REGION Network 15
   // ***************************************************************************************************************************************************
   // 
   // TC MAP SDC OUT Function Block FB118 - Maps Traffic Cop Zone motion Function blocks. Motion commands are determined at the zone position level and indexed by Zone number and stored in 
   //  "DB116_TC_ZoneMotionControl" DB. Block copies Traffic cop motion commands to the respective Carrier trafic cop and stores in TC_SDC_OUT Tag which is indexed by carrier number. 
   // 
   // ***************************************************************************************************************************************************
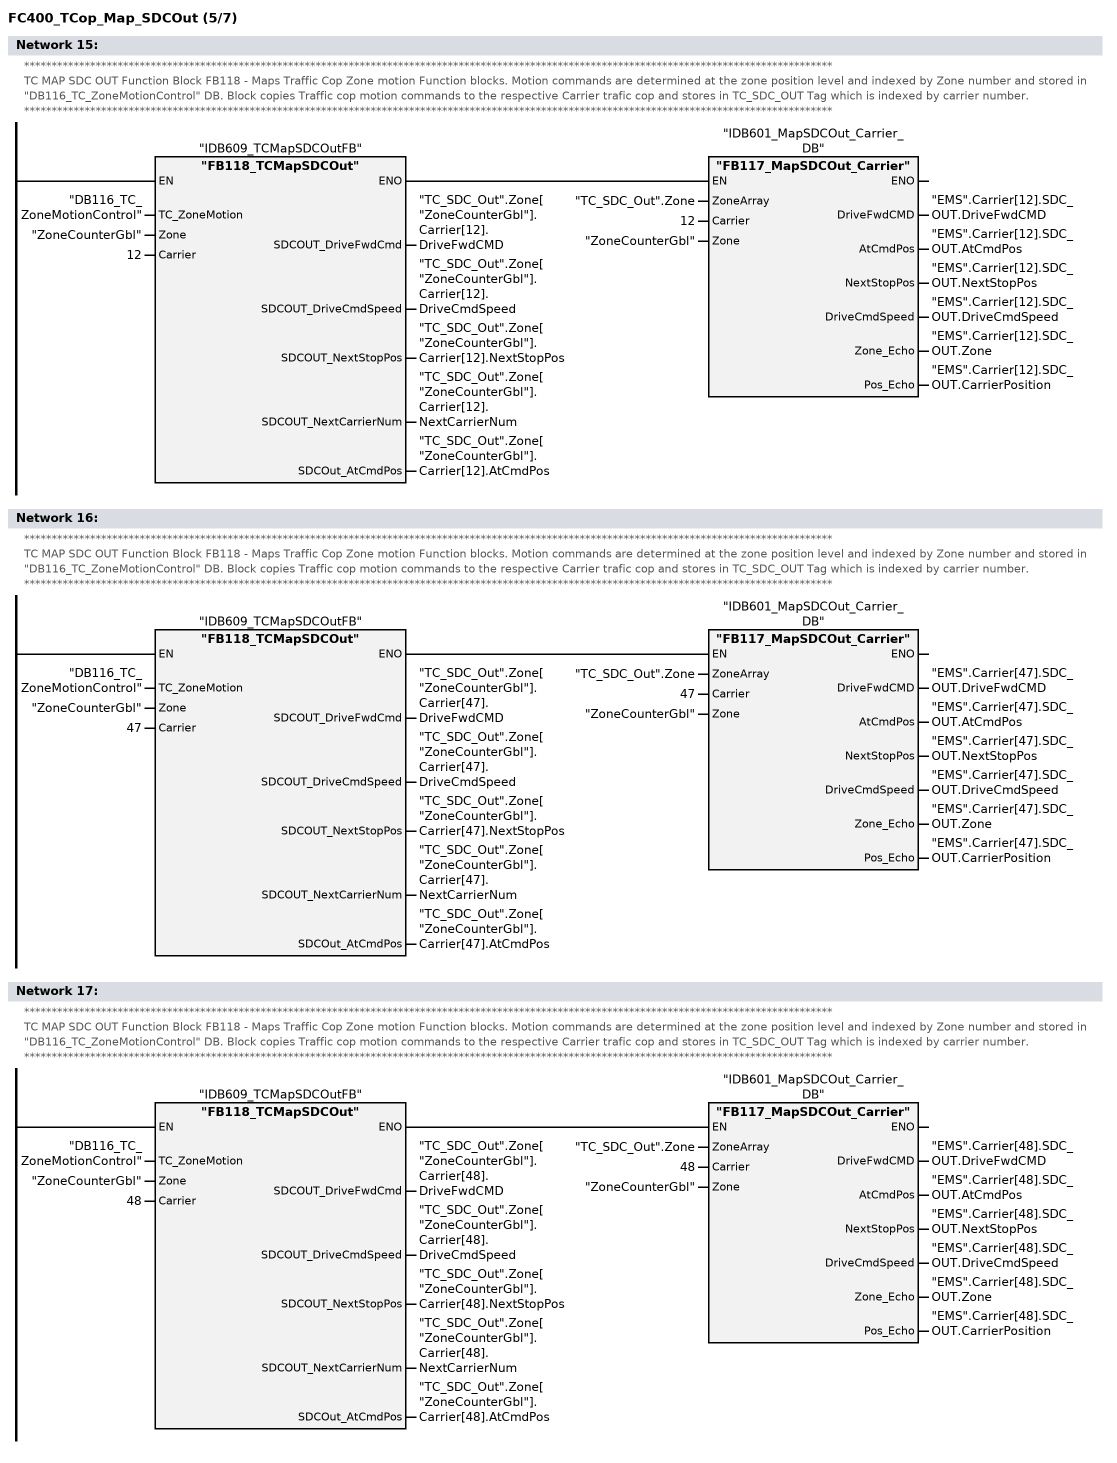
   RUNG wire#powerrail
      "IDB609_TCMapSDCOutFB"(TC_ZoneMotion := "DB116_TC_ZoneMotionControl", Zone := "ZoneCounterGbl", Carrier := 12, SDCOUT_DriveFwdCmd => "TC_SDC_Out".Zone["ZoneCounterGbl"].Carrier[12].DriveFwdCMD, SDCOUT_DriveCmdSpeed => "TC_SDC_Out".Zone["ZoneCounterGbl"].Carrier[12].DriveCmdSpeed, SDCOUT_NextStopPos => "TC_SDC_Out".Zone["ZoneCounterGbl"].Carrier[12].NextStopPos, SDCOUT_NextCarrierNum => "TC_SDC_Out".Zone["ZoneCounterGbl"].Carrier[12].NextCarrierNum, SDCOut_AtCmdPos => "TC_SDC_Out".Zone["ZoneCounterGbl"].Carrier[12].AtCmdPos)
      "IDB601_MapSDCOut_Carrier_DB"(ZoneArray := "TC_SDC_Out".Zone, Carrier := 12, Zone := "ZoneCounterGbl", DriveFwdCMD => "EMS".Carrier[12].SDC_OUT.DriveFwdCMD, AtCmdPos => "EMS".Carrier[12].SDC_OUT.AtCmdPos, NextStopPos => "EMS".Carrier[12].SDC_OUT.NextStopPos, DriveCmdSpeed => "EMS".Carrier[12].SDC_OUT.DriveCmdSpeed, Zone_Echo => "EMS".Carrier[12].SDC_OUT.Zone, Pos_Echo => "EMS".Carrier[12].SDC_OUT.CarrierPosition)
   END_RUNG
   // the same network as SCL:
   "IDB609_TCMapSDCOutFB"(TC_ZoneMotion := "DB116_TC_ZoneMotionControl",   // "FB118_TCMapSDCOut"
                          Zone := "ZoneCounterGbl",
                          Carrier := 12,
                          SDCOUT_DriveFwdCmd => "TC_SDC_Out".Zone["ZoneCounterGbl"].Carrier[12].DriveFwdCMD,
                          SDCOUT_DriveCmdSpeed => "TC_SDC_Out".Zone["ZoneCounterGbl"].Carrier[12].DriveCmdSpeed,
                          SDCOUT_NextStopPos => "TC_SDC_Out".Zone["ZoneCounterGbl"].Carrier[12].NextStopPos,
                          SDCOUT_NextCarrierNum => "TC_SDC_Out".Zone["ZoneCounterGbl"].Carrier[12].NextCarrierNum,
                          SDCOut_AtCmdPos => "TC_SDC_Out".Zone["ZoneCounterGbl"].Carrier[12].AtCmdPos,
                          ENO => #_w1);
   IF #_w1 THEN
       "IDB601_MapSDCOut_Carrier_DB"(ZoneArray := "TC_SDC_Out".Zone,   // "FB117_MapSDCOut_Carrier"
                               Carrier := 12,
                               Zone := "ZoneCounterGbl",
                               DriveFwdCMD => "EMS".Carrier[12].SDC_OUT.DriveFwdCMD,
                               AtCmdPos => "EMS".Carrier[12].SDC_OUT.AtCmdPos,
                               NextStopPos => "EMS".Carrier[12].SDC_OUT.NextStopPos,
                               DriveCmdSpeed => "EMS".Carrier[12].SDC_OUT.DriveCmdSpeed,
                               Zone_Echo => "EMS".Carrier[12].SDC_OUT.Zone,
                               Pos_Echo => "EMS".Carrier[12].SDC_OUT.CarrierPosition);
   END_IF;
END_REGION

REGION Network 16
   // ***************************************************************************************************************************************************
   // 
   // TC MAP SDC OUT Function Block FB118 - Maps Traffic Cop Zone motion Function blocks. Motion commands are determined at the zone position level and indexed by Zone number and stored in 
   //  "DB116_TC_ZoneMotionControl" DB. Block copies Traffic cop motion commands to the respective Carrier trafic cop and stores in TC_SDC_OUT Tag which is indexed by carrier number. 
   // 
   // ***************************************************************************************************************************************************
   RUNG wire#powerrail
      "IDB609_TCMapSDCOutFB"(TC_ZoneMotion := "DB116_TC_ZoneMotionControl", Zone := "ZoneCounterGbl", Carrier := 47, SDCOUT_DriveFwdCmd => "TC_SDC_Out".Zone["ZoneCounterGbl"].Carrier[47].DriveFwdCMD, SDCOUT_DriveCmdSpeed => "TC_SDC_Out".Zone["ZoneCounterGbl"].Carrier[47].DriveCmdSpeed, SDCOUT_NextStopPos => "TC_SDC_Out".Zone["ZoneCounterGbl"].Carrier[47].NextStopPos, SDCOUT_NextCarrierNum => "TC_SDC_Out".Zone["ZoneCounterGbl"].Carrier[47].NextCarrierNum, SDCOut_AtCmdPos => "TC_SDC_Out".Zone["ZoneCounterGbl"].Carrier[47].AtCmdPos)
      "IDB601_MapSDCOut_Carrier_DB"(ZoneArray := "TC_SDC_Out".Zone, Carrier := 47, Zone := "ZoneCounterGbl", DriveFwdCMD => "EMS".Carrier[47].SDC_OUT.DriveFwdCMD, AtCmdPos => "EMS".Carrier[47].SDC_OUT.AtCmdPos, NextStopPos => "EMS".Carrier[47].SDC_OUT.NextStopPos, DriveCmdSpeed => "EMS".Carrier[47].SDC_OUT.DriveCmdSpeed, Zone_Echo => "EMS".Carrier[47].SDC_OUT.Zone, Pos_Echo => "EMS".Carrier[47].SDC_OUT.CarrierPosition)
   END_RUNG
   // the same network as SCL:
   "IDB609_TCMapSDCOutFB"(TC_ZoneMotion := "DB116_TC_ZoneMotionControl",   // "FB118_TCMapSDCOut"
                          Zone := "ZoneCounterGbl",
                          Carrier := 47,
                          SDCOUT_DriveFwdCmd => "TC_SDC_Out".Zone["ZoneCounterGbl"].Carrier[47].DriveFwdCMD,
                          SDCOUT_DriveCmdSpeed => "TC_SDC_Out".Zone["ZoneCounterGbl"].Carrier[47].DriveCmdSpeed,
                          SDCOUT_NextStopPos => "TC_SDC_Out".Zone["ZoneCounterGbl"].Carrier[47].NextStopPos,
                          SDCOUT_NextCarrierNum => "TC_SDC_Out".Zone["ZoneCounterGbl"].Carrier[47].NextCarrierNum,
                          SDCOut_AtCmdPos => "TC_SDC_Out".Zone["ZoneCounterGbl"].Carrier[47].AtCmdPos,
                          ENO => #_w1);
   IF #_w1 THEN
       "IDB601_MapSDCOut_Carrier_DB"(ZoneArray := "TC_SDC_Out".Zone,   // "FB117_MapSDCOut_Carrier"
                               Carrier := 47,
                               Zone := "ZoneCounterGbl",
                               DriveFwdCMD => "EMS".Carrier[47].SDC_OUT.DriveFwdCMD,
                               AtCmdPos => "EMS".Carrier[47].SDC_OUT.AtCmdPos,
                               NextStopPos => "EMS".Carrier[47].SDC_OUT.NextStopPos,
                               DriveCmdSpeed => "EMS".Carrier[47].SDC_OUT.DriveCmdSpeed,
                               Zone_Echo => "EMS".Carrier[47].SDC_OUT.Zone,
                               Pos_Echo => "EMS".Carrier[47].SDC_OUT.CarrierPosition);
   END_IF;
END_REGION

REGION Network 17
   // ***************************************************************************************************************************************************
   // 
   // TC MAP SDC OUT Function Block FB118 - Maps Traffic Cop Zone motion Function blocks. Motion commands are determined at the zone position level and indexed by Zone number and stored in 
   //  "DB116_TC_ZoneMotionControl" DB. Block copies Traffic cop motion commands to the respective Carrier trafic cop and stores in TC_SDC_OUT Tag which is indexed by carrier number. 
   // 
   // ***************************************************************************************************************************************************
   RUNG wire#powerrail
      "IDB609_TCMapSDCOutFB"(TC_ZoneMotion := "DB116_TC_ZoneMotionControl", Zone := "ZoneCounterGbl", Carrier := 48, SDCOUT_DriveFwdCmd => "TC_SDC_Out".Zone["ZoneCounterGbl"].Carrier[48].DriveFwdCMD, SDCOUT_DriveCmdSpeed => "TC_SDC_Out".Zone["ZoneCounterGbl"].Carrier[48].DriveCmdSpeed, SDCOUT_NextStopPos => "TC_SDC_Out".Zone["ZoneCounterGbl"].Carrier[48].NextStopPos, SDCOUT_NextCarrierNum => "TC_SDC_Out".Zone["ZoneCounterGbl"].Carrier[48].NextCarrierNum, SDCOut_AtCmdPos => "TC_SDC_Out".Zone["ZoneCounterGbl"].Carrier[48].AtCmdPos)
      "IDB601_MapSDCOut_Carrier_DB"(ZoneArray := "TC_SDC_Out".Zone, Carrier := 48, Zone := "ZoneCounterGbl", DriveFwdCMD => "EMS".Carrier[48].SDC_OUT.DriveFwdCMD, AtCmdPos => "EMS".Carrier[48].SDC_OUT.AtCmdPos, NextStopPos => "EMS".Carrier[48].SDC_OUT.NextStopPos, DriveCmdSpeed => "EMS".Carrier[48].SDC_OUT.DriveCmdSpeed, Zone_Echo => "EMS".Carrier[48].SDC_OUT.Zone, Pos_Echo => "EMS".Carrier[48].SDC_OUT.CarrierPosition)
   END_RUNG
   // the same network as SCL:
   "IDB609_TCMapSDCOutFB"(TC_ZoneMotion := "DB116_TC_ZoneMotionControl",   // "FB118_TCMapSDCOut"
                          Zone := "ZoneCounterGbl",
                          Carrier := 48,
                          SDCOUT_DriveFwdCmd => "TC_SDC_Out".Zone["ZoneCounterGbl"].Carrier[48].DriveFwdCMD,
                          SDCOUT_DriveCmdSpeed => "TC_SDC_Out".Zone["ZoneCounterGbl"].Carrier[48].DriveCmdSpeed,
                          SDCOUT_NextStopPos => "TC_SDC_Out".Zone["ZoneCounterGbl"].Carrier[48].NextStopPos,
                          SDCOUT_NextCarrierNum => "TC_SDC_Out".Zone["ZoneCounterGbl"].Carrier[48].NextCarrierNum,
                          SDCOut_AtCmdPos => "TC_SDC_Out".Zone["ZoneCounterGbl"].Carrier[48].AtCmdPos,
                          ENO => #_w1);
   IF #_w1 THEN
       "IDB601_MapSDCOut_Carrier_DB"(ZoneArray := "TC_SDC_Out".Zone,   // "FB117_MapSDCOut_Carrier"
                               Carrier := 48,
                               Zone := "ZoneCounterGbl",
                               DriveFwdCMD => "EMS".Carrier[48].SDC_OUT.DriveFwdCMD,
                               AtCmdPos => "EMS".Carrier[48].SDC_OUT.AtCmdPos,
                               NextStopPos => "EMS".Carrier[48].SDC_OUT.NextStopPos,
                               DriveCmdSpeed => "EMS".Carrier[48].SDC_OUT.DriveCmdSpeed,
                               Zone_Echo => "EMS".Carrier[48].SDC_OUT.Zone,
                               Pos_Echo => "EMS".Carrier[48].SDC_OUT.CarrierPosition);
   END_IF;
END_REGION

REGION Network 18
   // ***************************************************************************************************************************************************
   // 
   // TC MAP SDC OUT Function Block FB118 - Maps Traffic Cop Zone motion Function blocks. Motion commands are determined at the zone position level and indexed by Zone number and stored in 
   //  "DB116_TC_ZoneMotionControl" DB. Block copies Traffic cop motion commands to the respective Carrier trafic cop and stores in TC_SDC_OUT Tag which is indexed by carrier number. 
   // 
   // ***************************************************************************************************************************************************
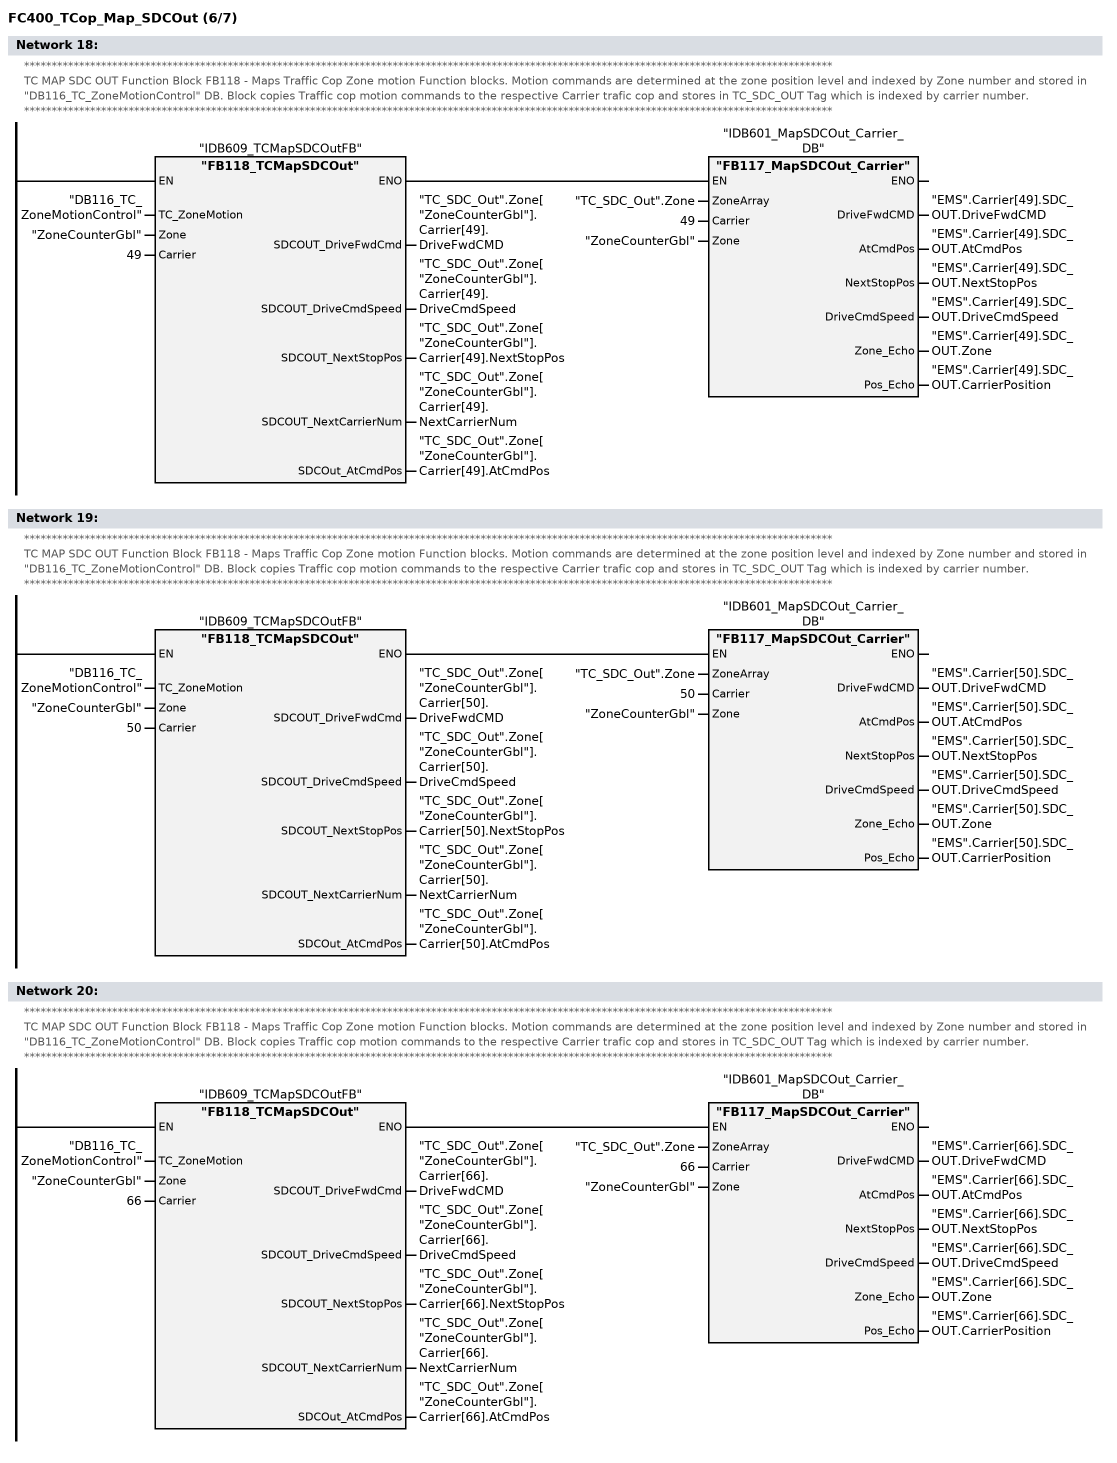
   RUNG wire#powerrail
      "IDB609_TCMapSDCOutFB"(TC_ZoneMotion := "DB116_TC_ZoneMotionControl", Zone := "ZoneCounterGbl", Carrier := 49, SDCOUT_DriveFwdCmd => "TC_SDC_Out".Zone["ZoneCounterGbl"].Carrier[49].DriveFwdCMD, SDCOUT_DriveCmdSpeed => "TC_SDC_Out".Zone["ZoneCounterGbl"].Carrier[49].DriveCmdSpeed, SDCOUT_NextStopPos => "TC_SDC_Out".Zone["ZoneCounterGbl"].Carrier[49].NextStopPos, SDCOUT_NextCarrierNum => "TC_SDC_Out".Zone["ZoneCounterGbl"].Carrier[49].NextCarrierNum, SDCOut_AtCmdPos => "TC_SDC_Out".Zone["ZoneCounterGbl"].Carrier[49].AtCmdPos)
      "IDB601_MapSDCOut_Carrier_DB"(ZoneArray := "TC_SDC_Out".Zone, Carrier := 49, Zone := "ZoneCounterGbl", DriveFwdCMD => "EMS".Carrier[49].SDC_OUT.DriveFwdCMD, AtCmdPos => "EMS".Carrier[49].SDC_OUT.AtCmdPos, NextStopPos => "EMS".Carrier[49].SDC_OUT.NextStopPos, DriveCmdSpeed => "EMS".Carrier[49].SDC_OUT.DriveCmdSpeed, Zone_Echo => "EMS".Carrier[49].SDC_OUT.Zone, Pos_Echo => "EMS".Carrier[49].SDC_OUT.CarrierPosition)
   END_RUNG
   // the same network as SCL:
   "IDB609_TCMapSDCOutFB"(TC_ZoneMotion := "DB116_TC_ZoneMotionControl",   // "FB118_TCMapSDCOut"
                          Zone := "ZoneCounterGbl",
                          Carrier := 49,
                          SDCOUT_DriveFwdCmd => "TC_SDC_Out".Zone["ZoneCounterGbl"].Carrier[49].DriveFwdCMD,
                          SDCOUT_DriveCmdSpeed => "TC_SDC_Out".Zone["ZoneCounterGbl"].Carrier[49].DriveCmdSpeed,
                          SDCOUT_NextStopPos => "TC_SDC_Out".Zone["ZoneCounterGbl"].Carrier[49].NextStopPos,
                          SDCOUT_NextCarrierNum => "TC_SDC_Out".Zone["ZoneCounterGbl"].Carrier[49].NextCarrierNum,
                          SDCOut_AtCmdPos => "TC_SDC_Out".Zone["ZoneCounterGbl"].Carrier[49].AtCmdPos,
                          ENO => #_w1);
   IF #_w1 THEN
       "IDB601_MapSDCOut_Carrier_DB"(ZoneArray := "TC_SDC_Out".Zone,   // "FB117_MapSDCOut_Carrier"
                               Carrier := 49,
                               Zone := "ZoneCounterGbl",
                               DriveFwdCMD => "EMS".Carrier[49].SDC_OUT.DriveFwdCMD,
                               AtCmdPos => "EMS".Carrier[49].SDC_OUT.AtCmdPos,
                               NextStopPos => "EMS".Carrier[49].SDC_OUT.NextStopPos,
                               DriveCmdSpeed => "EMS".Carrier[49].SDC_OUT.DriveCmdSpeed,
                               Zone_Echo => "EMS".Carrier[49].SDC_OUT.Zone,
                               Pos_Echo => "EMS".Carrier[49].SDC_OUT.CarrierPosition);
   END_IF;
END_REGION

REGION Network 19
   // ***************************************************************************************************************************************************
   // 
   // TC MAP SDC OUT Function Block FB118 - Maps Traffic Cop Zone motion Function blocks. Motion commands are determined at the zone position level and indexed by Zone number and stored in 
   //  "DB116_TC_ZoneMotionControl" DB. Block copies Traffic cop motion commands to the respective Carrier trafic cop and stores in TC_SDC_OUT Tag which is indexed by carrier number. 
   // 
   // ***************************************************************************************************************************************************
   RUNG wire#powerrail
      "IDB609_TCMapSDCOutFB"(TC_ZoneMotion := "DB116_TC_ZoneMotionControl", Zone := "ZoneCounterGbl", Carrier := 50, SDCOUT_DriveFwdCmd => "TC_SDC_Out".Zone["ZoneCounterGbl"].Carrier[50].DriveFwdCMD, SDCOUT_DriveCmdSpeed => "TC_SDC_Out".Zone["ZoneCounterGbl"].Carrier[50].DriveCmdSpeed, SDCOUT_NextStopPos => "TC_SDC_Out".Zone["ZoneCounterGbl"].Carrier[50].NextStopPos, SDCOUT_NextCarrierNum => "TC_SDC_Out".Zone["ZoneCounterGbl"].Carrier[50].NextCarrierNum, SDCOut_AtCmdPos => "TC_SDC_Out".Zone["ZoneCounterGbl"].Carrier[50].AtCmdPos)
      "IDB601_MapSDCOut_Carrier_DB"(ZoneArray := "TC_SDC_Out".Zone, Carrier := 50, Zone := "ZoneCounterGbl", DriveFwdCMD => "EMS".Carrier[50].SDC_OUT.DriveFwdCMD, AtCmdPos => "EMS".Carrier[50].SDC_OUT.AtCmdPos, NextStopPos => "EMS".Carrier[50].SDC_OUT.NextStopPos, DriveCmdSpeed => "EMS".Carrier[50].SDC_OUT.DriveCmdSpeed, Zone_Echo => "EMS".Carrier[50].SDC_OUT.Zone, Pos_Echo => "EMS".Carrier[50].SDC_OUT.CarrierPosition)
   END_RUNG
   // the same network as SCL:
   "IDB609_TCMapSDCOutFB"(TC_ZoneMotion := "DB116_TC_ZoneMotionControl",   // "FB118_TCMapSDCOut"
                          Zone := "ZoneCounterGbl",
                          Carrier := 50,
                          SDCOUT_DriveFwdCmd => "TC_SDC_Out".Zone["ZoneCounterGbl"].Carrier[50].DriveFwdCMD,
                          SDCOUT_DriveCmdSpeed => "TC_SDC_Out".Zone["ZoneCounterGbl"].Carrier[50].DriveCmdSpeed,
                          SDCOUT_NextStopPos => "TC_SDC_Out".Zone["ZoneCounterGbl"].Carrier[50].NextStopPos,
                          SDCOUT_NextCarrierNum => "TC_SDC_Out".Zone["ZoneCounterGbl"].Carrier[50].NextCarrierNum,
                          SDCOut_AtCmdPos => "TC_SDC_Out".Zone["ZoneCounterGbl"].Carrier[50].AtCmdPos,
                          ENO => #_w1);
   IF #_w1 THEN
       "IDB601_MapSDCOut_Carrier_DB"(ZoneArray := "TC_SDC_Out".Zone,   // "FB117_MapSDCOut_Carrier"
                               Carrier := 50,
                               Zone := "ZoneCounterGbl",
                               DriveFwdCMD => "EMS".Carrier[50].SDC_OUT.DriveFwdCMD,
                               AtCmdPos => "EMS".Carrier[50].SDC_OUT.AtCmdPos,
                               NextStopPos => "EMS".Carrier[50].SDC_OUT.NextStopPos,
                               DriveCmdSpeed => "EMS".Carrier[50].SDC_OUT.DriveCmdSpeed,
                               Zone_Echo => "EMS".Carrier[50].SDC_OUT.Zone,
                               Pos_Echo => "EMS".Carrier[50].SDC_OUT.CarrierPosition);
   END_IF;
END_REGION

REGION Network 20
   // ***************************************************************************************************************************************************
   // 
   // TC MAP SDC OUT Function Block FB118 - Maps Traffic Cop Zone motion Function blocks. Motion commands are determined at the zone position level and indexed by Zone number and stored in 
   //  "DB116_TC_ZoneMotionControl" DB. Block copies Traffic cop motion commands to the respective Carrier trafic cop and stores in TC_SDC_OUT Tag which is indexed by carrier number. 
   // 
   // ***************************************************************************************************************************************************
   RUNG wire#powerrail
      "IDB609_TCMapSDCOutFB"(TC_ZoneMotion := "DB116_TC_ZoneMotionControl", Zone := "ZoneCounterGbl", Carrier := 66, SDCOUT_DriveFwdCmd => "TC_SDC_Out".Zone["ZoneCounterGbl"].Carrier[66].DriveFwdCMD, SDCOUT_DriveCmdSpeed => "TC_SDC_Out".Zone["ZoneCounterGbl"].Carrier[66].DriveCmdSpeed, SDCOUT_NextStopPos => "TC_SDC_Out".Zone["ZoneCounterGbl"].Carrier[66].NextStopPos, SDCOUT_NextCarrierNum => "TC_SDC_Out".Zone["ZoneCounterGbl"].Carrier[66].NextCarrierNum, SDCOut_AtCmdPos => "TC_SDC_Out".Zone["ZoneCounterGbl"].Carrier[66].AtCmdPos)
      "IDB601_MapSDCOut_Carrier_DB"(ZoneArray := "TC_SDC_Out".Zone, Carrier := 66, Zone := "ZoneCounterGbl", DriveFwdCMD => "EMS".Carrier[66].SDC_OUT.DriveFwdCMD, AtCmdPos => "EMS".Carrier[66].SDC_OUT.AtCmdPos, NextStopPos => "EMS".Carrier[66].SDC_OUT.NextStopPos, DriveCmdSpeed => "EMS".Carrier[66].SDC_OUT.DriveCmdSpeed, Zone_Echo => "EMS".Carrier[66].SDC_OUT.Zone, Pos_Echo => "EMS".Carrier[66].SDC_OUT.CarrierPosition)
   END_RUNG
   // the same network as SCL:
   "IDB609_TCMapSDCOutFB"(TC_ZoneMotion := "DB116_TC_ZoneMotionControl",   // "FB118_TCMapSDCOut"
                          Zone := "ZoneCounterGbl",
                          Carrier := 66,
                          SDCOUT_DriveFwdCmd => "TC_SDC_Out".Zone["ZoneCounterGbl"].Carrier[66].DriveFwdCMD,
                          SDCOUT_DriveCmdSpeed => "TC_SDC_Out".Zone["ZoneCounterGbl"].Carrier[66].DriveCmdSpeed,
                          SDCOUT_NextStopPos => "TC_SDC_Out".Zone["ZoneCounterGbl"].Carrier[66].NextStopPos,
                          SDCOUT_NextCarrierNum => "TC_SDC_Out".Zone["ZoneCounterGbl"].Carrier[66].NextCarrierNum,
                          SDCOut_AtCmdPos => "TC_SDC_Out".Zone["ZoneCounterGbl"].Carrier[66].AtCmdPos,
                          ENO => #_w1);
   IF #_w1 THEN
       "IDB601_MapSDCOut_Carrier_DB"(ZoneArray := "TC_SDC_Out".Zone,   // "FB117_MapSDCOut_Carrier"
                               Carrier := 66,
                               Zone := "ZoneCounterGbl",
                               DriveFwdCMD => "EMS".Carrier[66].SDC_OUT.DriveFwdCMD,
                               AtCmdPos => "EMS".Carrier[66].SDC_OUT.AtCmdPos,
                               NextStopPos => "EMS".Carrier[66].SDC_OUT.NextStopPos,
                               DriveCmdSpeed => "EMS".Carrier[66].SDC_OUT.DriveCmdSpeed,
                               Zone_Echo => "EMS".Carrier[66].SDC_OUT.Zone,
                               Pos_Echo => "EMS".Carrier[66].SDC_OUT.CarrierPosition);
   END_IF;
END_REGION

REGION Network 21
   // *********************************************************************************************************************************
   // 
   // Zone Index Counter - Used to Index  Zone Traffic Cop Carrier Information determined by the Zone Traffic cop FC  
   // 
   // **********************************************************************************************************************************
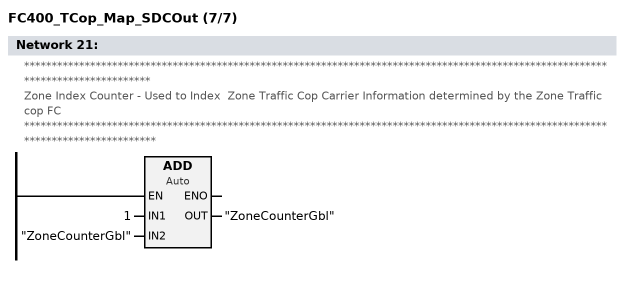
   RUNG wire#powerrail
      Add(in1 := 1, in2 := "ZoneCounterGbl", out => "ZoneCounterGbl")
   END_RUNG
   // the same network as SCL:
   "ZoneCounterGbl" := 1 + "ZoneCounterGbl";
END_REGION
END_FUNCTION

FUNCTION "FC500_FAULTS" : Void   // FC500, LAD
{ S7_Optimized_Access := 'TRUE' }
VERSION : 0.1
BEGIN

REGION Network 1
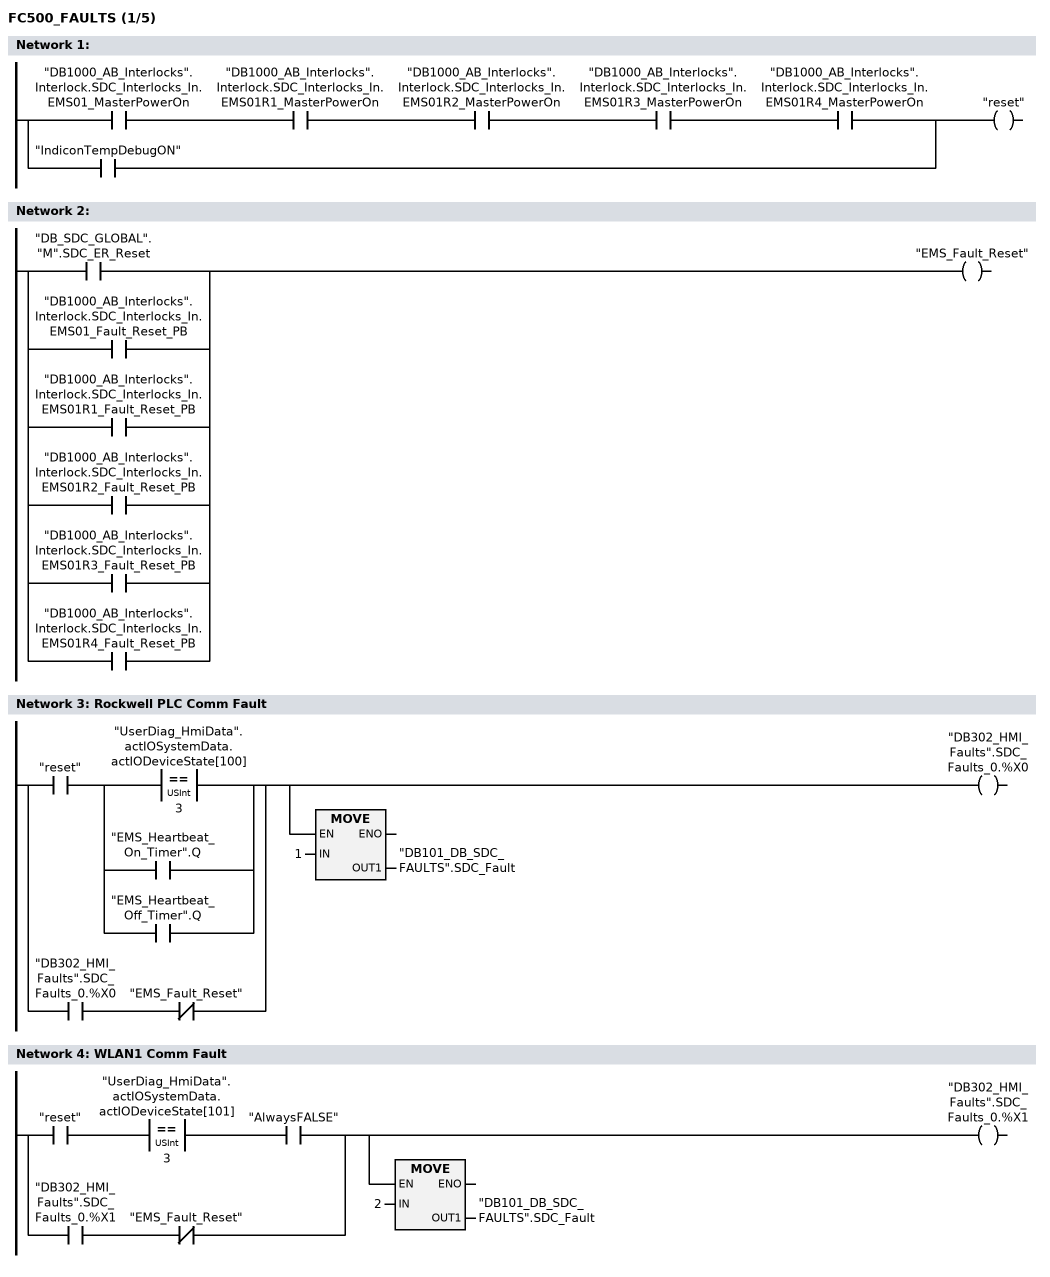
   RUNG wire#powerrail
      Contact( "DB1000_AB_Interlocks".Interlock.SDC_Interlocks_In.EMS01_MasterPowerOn )
      Contact( "DB1000_AB_Interlocks".Interlock.SDC_Interlocks_In.EMS01R1_MasterPowerOn )
      Contact( "DB1000_AB_Interlocks".Interlock.SDC_Interlocks_In.EMS01R2_MasterPowerOn )
      Contact( "DB1000_AB_Interlocks".Interlock.SDC_Interlocks_In.EMS01R3_MasterPowerOn )
      Contact( "DB1000_AB_Interlocks".Interlock.SDC_Interlocks_In.EMS01R4_MasterPowerOn )
      wire#w1
      Coil( "reset" )
   END_RUNG
   RUNG wire#powerrail
      Contact( "IndiconTempDebugON" )
   END_RUNG wire#w1
   // the same network as SCL:
   "reset" := ("DB1000_AB_Interlocks".Interlock.SDC_Interlocks_In.EMS01_MasterPowerOn AND "DB1000_AB_Interlocks".Interlock.SDC_Interlocks_In.EMS01R1_MasterPowerOn AND "DB1000_AB_Interlocks".Interlock.SDC_Interlocks_In.EMS01R2_MasterPowerOn AND "DB1000_AB_Interlocks".Interlock.SDC_Interlocks_In.EMS01R3_MasterPowerOn AND "DB1000_AB_Interlocks".Interlock.SDC_Interlocks_In.EMS01R4_MasterPowerOn) OR "IndiconTempDebugON";
END_REGION

REGION Network 2
   RUNG wire#powerrail
      Contact( "DB_SDC_GLOBAL"."M".SDC_ER_Reset )
      wire#w1
      Coil( "EMS_Fault_Reset" )
   END_RUNG
   RUNG wire#powerrail
      Contact( "DB1000_AB_Interlocks".Interlock.SDC_Interlocks_In.EMS01_Fault_Reset_PB )
   END_RUNG wire#w1
   RUNG wire#powerrail
      Contact( "DB1000_AB_Interlocks".Interlock.SDC_Interlocks_In.EMS01R1_Fault_Reset_PB )
   END_RUNG wire#w1
   RUNG wire#powerrail
      Contact( "DB1000_AB_Interlocks".Interlock.SDC_Interlocks_In.EMS01R2_Fault_Reset_PB )
   END_RUNG wire#w1
   RUNG wire#powerrail
      Contact( "DB1000_AB_Interlocks".Interlock.SDC_Interlocks_In.EMS01R3_Fault_Reset_PB )
   END_RUNG wire#w1
   RUNG wire#powerrail
      Contact( "DB1000_AB_Interlocks".Interlock.SDC_Interlocks_In.EMS01R4_Fault_Reset_PB )
   END_RUNG wire#w1
   // the same network as SCL:
   "EMS_Fault_Reset" := "DB_SDC_GLOBAL"."M".SDC_ER_Reset OR "DB1000_AB_Interlocks".Interlock.SDC_Interlocks_In.EMS01_Fault_Reset_PB OR "DB1000_AB_Interlocks".Interlock.SDC_Interlocks_In.EMS01R1_Fault_Reset_PB OR "DB1000_AB_Interlocks".Interlock.SDC_Interlocks_In.EMS01R2_Fault_Reset_PB OR "DB1000_AB_Interlocks".Interlock.SDC_Interlocks_In.EMS01R3_Fault_Reset_PB OR "DB1000_AB_Interlocks".Interlock.SDC_Interlocks_In.EMS01R4_Fault_Reset_PB;
END_REGION

REGION Network 3: Rockwell PLC Comm Fault
   RUNG wire#powerrail
      Contact( "reset" )
      wire#w1
      { S7_Templates := "SrcType := USInt" } EQ_Contact(in1 := "UserDiag_HmiData".actIOSystemData.actIODeviceState[100], in2 := 3)
      wire#w2
      Coil( "DB302_HMI_Faults".SDC_Faults_0.%X0 )
   END_RUNG
   RUNG wire#w1
      Contact( "EMS_Heartbeat_On_Timer".Q )
   END_RUNG wire#w2
   RUNG wire#w1
      Contact( "EMS_Heartbeat_Off_Timer".Q )
   END_RUNG wire#w2
   RUNG wire#powerrail
      Contact( "DB302_HMI_Faults".SDC_Faults_0.%X0 )
      I_Contact( "EMS_Fault_Reset" )
   END_RUNG wire#w2
   RUNG wire#w2
      Move(in := 1, out1 => "DB101_DB_SDC_FAULTS".SDC_Fault)
   END_RUNG
   // the same network as SCL:
   "DB302_HMI_Faults".SDC_Faults_0.%X0 := ("reset" AND (("UserDiag_HmiData".actIOSystemData.actIODeviceState[100] = 3) OR "EMS_Heartbeat_On_Timer".Q OR "EMS_Heartbeat_Off_Timer".Q)) OR ("DB302_HMI_Faults".SDC_Faults_0.%X0 AND NOT "EMS_Fault_Reset");
   IF "DB302_HMI_Faults".SDC_Faults_0.%X0 THEN "DB101_DB_SDC_FAULTS".SDC_Fault := 1; END_IF;
END_REGION

REGION Network 4: WLAN1 Comm Fault
   RUNG wire#powerrail
      Contact( "reset" )
      { S7_Templates := "SrcType := USInt" } EQ_Contact(in1 := "UserDiag_HmiData".actIOSystemData.actIODeviceState[101], in2 := 3)
      Contact( "AlwaysFALSE" )
      wire#w1
      Coil( "DB302_HMI_Faults".SDC_Faults_0.%X1 )
   END_RUNG
   RUNG wire#powerrail
      Contact( "DB302_HMI_Faults".SDC_Faults_0.%X1 )
      I_Contact( "EMS_Fault_Reset" )
   END_RUNG wire#w1
   RUNG wire#w1
      Move(in := 2, out1 => "DB101_DB_SDC_FAULTS".SDC_Fault)
   END_RUNG
   // the same network as SCL:
   "DB302_HMI_Faults".SDC_Faults_0.%X1 := ("reset" AND ("UserDiag_HmiData".actIOSystemData.actIODeviceState[101] = 3) AND "AlwaysFALSE") OR ("DB302_HMI_Faults".SDC_Faults_0.%X1 AND NOT "EMS_Fault_Reset");
   IF "DB302_HMI_Faults".SDC_Faults_0.%X1 THEN "DB101_DB_SDC_FAULTS".SDC_Fault := 2; END_IF;
END_REGION

REGION Network 5: WLAN2 Comm Fault